(* Logix 5000 project; controller MV vendor 1 type 14 code 217 rev 31.11; software revision 31.00; part 25 of 53 *)
(* tags used below, declared in another part *)
   Alarm_Reset : BOOL;
   comms_to_blunger_write_enabled : BOOL;
   comms_to_fv_route_write_enabled : BOOL;
   comms_to_mv_route_write_enabled : BOOL;
   CWD : CHECKWORD_FLAGS;
   Default_Check_Time : DINT;
   fvrroute_slc_still_active : BOOL;
   Item_Faults_Are_Latched : BOOL;
   Item_Simulation_Flag : BOOL;
   MC_CH2_FM_AI : PlantItem;   // CH2_FM
   mc_comms_from_brewhouse : MESSAGE;
   mc_comms_from_brewhouse_timer : TIMER;
   mc_comms_to_blunger : MESSAGE;
   mc_comms_to_blunger_timer : TIMER;
   mc_comms_to_fv_route : MESSAGE;
   mc_comms_to_fv_route_timer : TIMER;
   mc_comms_to_mv_route : MESSAGE;
   mc_comms_to_mv_route_timer : TIMER;
   MC_N23 : INT[255];   // P2 FLOW Control block and da ta for P2 flowrate P ID loop
   MC_P1 : PlantItem;   // P1
   MC_P1_ALARM : ALARM_DIGITAL;
   MC_P1_D : ALIAS FOR RIO_Rack_2:10:O.Data.0;
   MC_P1_R : ALIAS FOR RIO_Rack_2:11:I.Data.0;
   MC_P1_T : ALIAS FOR RIO_Rack_2:11:I.Data.15;
   MC_P2 : PlantItem;   // P2
   MC_P2_ALARM : ALARM_DIGITAL;
   MC_P2_D : ALIAS FOR RIO_Rack_2:10:O.Data.1;
   MC_P2_Flow_PID : PID;
   MC_P2_R : ALIAS FOR RIO_Rack_2:11:I.Data.1;
   MC_P2_T : ALIAS FOR RIO_Rack_2:11:I.Data.16;
   MC_P3 : PlantItem;   // P3
   MC_P3_ALARM : ALARM_DIGITAL;
   MC_P3_D : ALIAS FOR RIO_Rack_2:10:O.Data.2;
   MC_P3_R : ALIAS FOR RIO_Rack_2:11:I.Data.2;
   MC_P4 : PlantItem;   // P4
   MC_P4_ALARM : ALARM_DIGITAL;
   MC_P4_D : ALIAS FOR RIO_Rack_2:10:O.Data.3;
   MC_P4_R : ALIAS FOR RIO_Rack_2:11:I.Data.3;
   MC_SP_R1_1 : PlantItem;   // SP_R1_1
   MC_SP_R1_1_ALARM : ALARM_DIGITAL;
   MC_SP_R1_1_D : ALIAS FOR RIO_Rack_2:10:O.Data.4;
   MC_SP_R1_1_R : ALIAS FOR RIO_Rack_2:11:I.Data.4;
   MC_SP_R2_1 : PlantItem;   // SP_R2_1
   MC_SP_R2_1_ALARM : ALARM_DIGITAL;
   MC_SP_R2_1_D : ALIAS FOR RIO_Rack_2:10:O.Data.5;
   MC_SP_R2_1_R : ALIAS FOR RIO_Rack_2:11:I.Data.5;
   MC_SP_R2_2 : PlantItem;   // SP_R2_2
   MC_SP_R2_2_ALARM : ALARM_DIGITAL;
   MC_SP_R2_2_D : ALIAS FOR RIO_Rack_2:10:O.Data.15;
   MC_SP_R2_2_R : ALIAS FOR RIO_Rack_2:11:I.Data.14;
   MC_SP_R3_1 : PlantItem;   // SP_R3_1
   MC_SP_R3_1_ALARM : ALARM_DIGITAL;
   MC_SP_R3_1_D : ALIAS FOR RIO_Rack_2:10:O.Data.6;
   MC_SP_R3_1_R : ALIAS FOR RIO_Rack_2:11:I.Data.6;
   MC_SP_R5_1 : PlantItem;   // SP_R5_1
   MC_SP_R5_1_ALARM : ALARM_DIGITAL;
   MC_SP_R5_1_D : ALIAS FOR RIO_Rack_2:10:O.Data.7;
   MC_SP_R5_1_R : ALIAS FOR RIO_Rack_2:11:I.Data.7;
   MC_SP_R5_2 : PlantItem;   // SP_R5_2
   MC_SP_R5_2_ALARM : ALARM_DIGITAL;
   MC_SP_R5_2_D : ALIAS FOR RIO_Rack_2:10:O.Data.8;
   MC_SP_R5_2_R : ALIAS FOR RIO_Rack_2:11:I.Data.8;
   MC_SP_R6_1 : PlantItem;   // SP_R6_1
   MC_SP_R6_1_ALARM : ALARM_DIGITAL;
   MC_SP_R6_1_D : ALIAS FOR RIO_Rack_2:10:O.Data.9;
   MC_SP_R6_1_R : ALIAS FOR RIO_Rack_2:11:I.Data.9;
   MC_SP_R6_2 : PlantItem;   // SP_R6_2
   MC_SP_R6_2_ALARM : ALARM_DIGITAL;
   MC_SP_R6_2_D : ALIAS FOR RIO_Rack_2:10:O.Data.10;
   MC_SP_R6_2_R : ALIAS FOR RIO_Rack_2:11:I.Data.10;
   MC_SP_R6_3 : PlantItem;   // SP_R6_3
   MC_SP_R6_3_ALARM : ALARM_DIGITAL;
   MC_SP_R6_3_D : ALIAS FOR RIO_Rack_2:10:O.Data.11;
   MC_SP_R6_3_R : ALIAS FOR RIO_Rack_2:11:I.Data.11;
   MC_SP_R6_4 : PlantItem;   // SP_R6_4
   MC_SP_R6_4_ALARM : ALARM_DIGITAL;
   MC_SP_R6_4_D : ALIAS FOR RIO_Rack_2:10:O.Data.12;
   MC_SP_R6_4_R : ALIAS FOR RIO_Rack_2:11:I.Data.12;
   MC_SP_R6_5 : PlantItem;   // SP_R6_5
   MC_SP_R6_5_ALARM : ALARM_DIGITAL;
   MC_SP_R6_5_D : ALIAS FOR RIO_Rack_2:10:O.Data.13;
   MC_SP_R6_5_R : ALIAS FOR RIO_Rack_2:11:I.Data.13;
   One_Second_One_Scan : ALIAS FOR One_Second_1_scan;
   reset_msg_interval : BOOL;
   Scada_Pump_Fault_No : DINT;
   Scada_Pump_H_Fault_No : DINT;
   Scada_Pump_T_Fault_No : DINT;
   Unused_Healthy_Feedback : BOOL;
   Unused_NotTripped_Feedback : BOOL;
(* MC_Common, continued *)

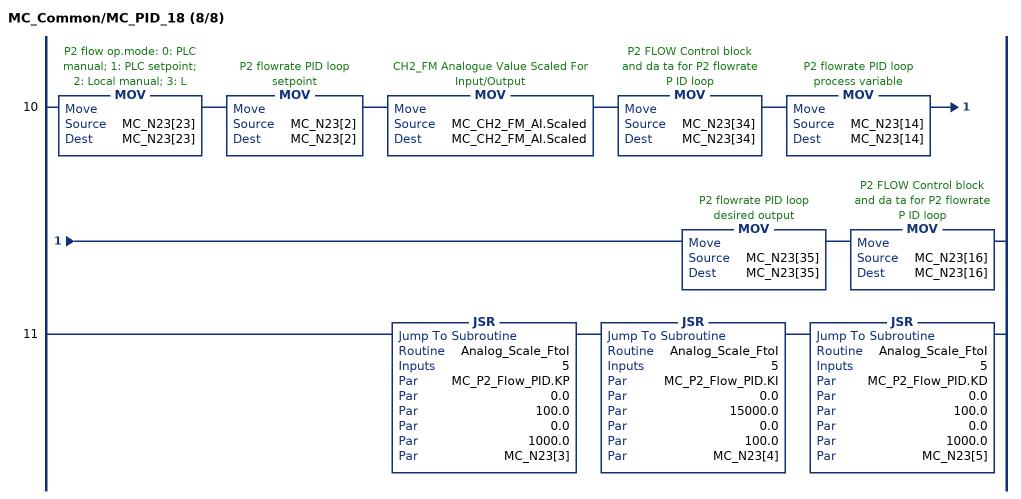
   [picture p462: MC_Common/MC_PID_18 rungs 10-11]
   10: MOV(MC_N23[23],MC_N23[23])MOV(MC_N23[2],MC_N23[2])MOV(MC_CH2_FM_AI.Scaled,MC_CH2_FM_AI.Scaled)MOV(MC_N23[34],MC_N23[34])MOV(MC_N23[14],MC_N23[14])MOV(MC_N23[35],MC_N23[35])MOV(MC_N23[16],MC_N23[16]);
   11: JSR(Analog_Scale_FtoI,5,MC_P2_Flow_PID.KP,0.0,100.0,0.0,1000.0,MC_N23[3])JSR(Analog_Scale_FtoI,5,MC_P2_Flow_PID.KI,0.0,15000.0,0.0,100.0,MC_N23[4])JSR(Analog_Scale_FtoI,5,MC_P2_Flow_PID.KD,0.0,100.0,0.0,1000.0,MC_N23[5]);
END_ROUTINE

ROUTINE MC_PLC_WRITE_REPLACEMENTS   (* ladder *)
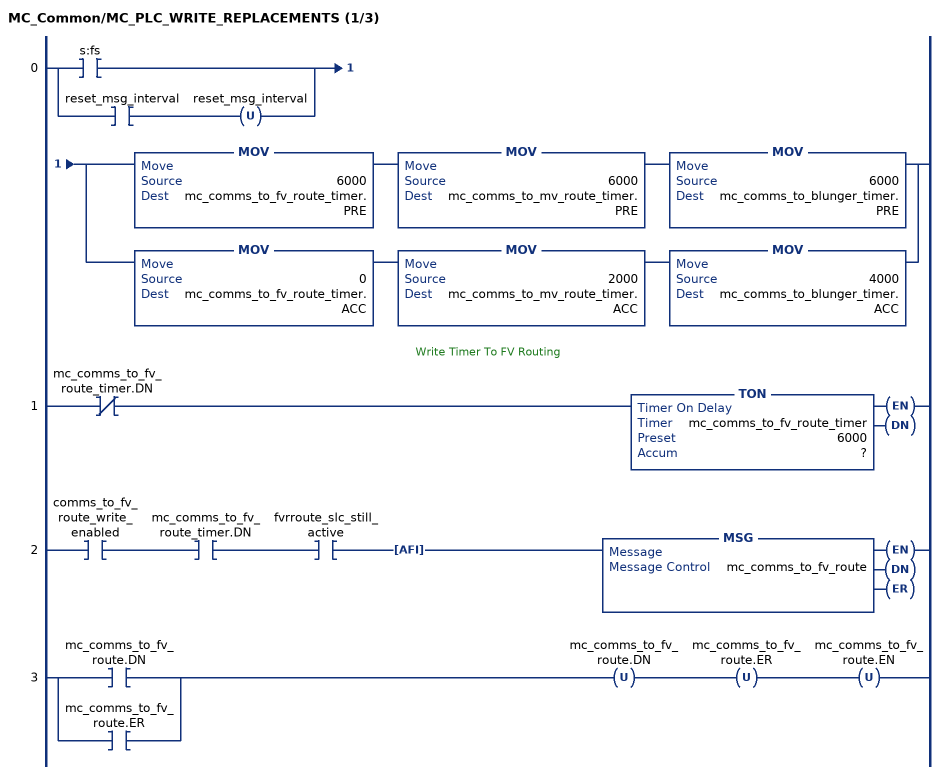
   0: [XIC(s:fs) ,XIC(reset_msg_interval) OTU(reset_msg_interval) ][MOV(6000,mc_comms_to_fv_route_timer.PRE) MOV(6000,mc_comms_to_mv_route_timer.PRE) MOV(6000,mc_comms_to_blunger_timer.PRE) ,MOV(0,mc_comms_to_fv_route_timer.ACC) MOV(2000,mc_comms_to_mv_route_timer.ACC) MOV(4000,mc_comms_to_blunger_timer.ACC) ];
   // Write Timer To FV Routing
   1: XIO(mc_comms_to_fv_route_timer.DN)TON(mc_comms_to_fv_route_timer,?,?);
   2: XIC(comms_to_fv_route_write_enabled)XIC(mc_comms_to_fv_route_timer.DN)XIC(fvrroute_slc_still_active)AFI()MSG(mc_comms_to_fv_route);
   3: [XIC(mc_comms_to_fv_route.DN) ,XIC(mc_comms_to_fv_route.ER) ]OTU(mc_comms_to_fv_route.DN)OTU(mc_comms_to_fv_route.ER)OTU(mc_comms_to_fv_route.EN);
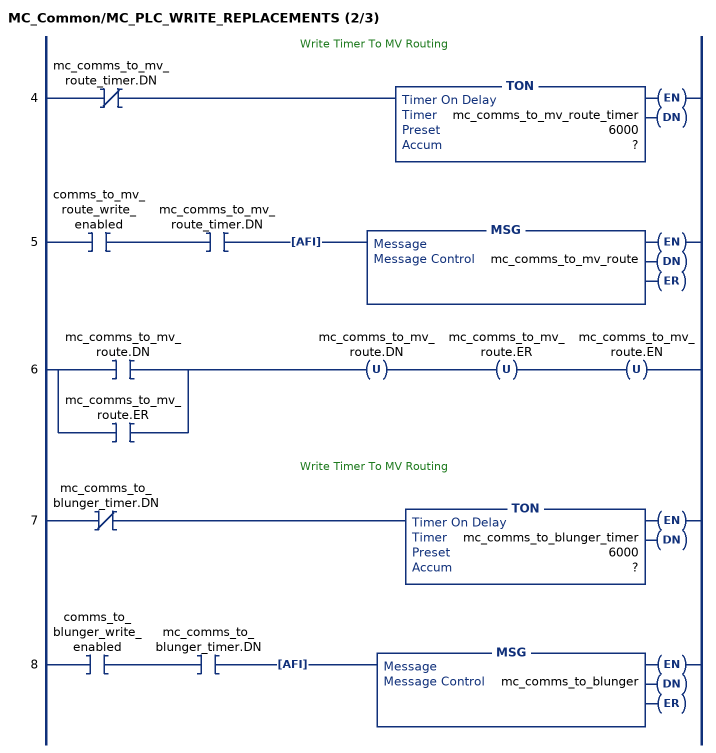
   // Write Timer To MV Routing
   4: XIO(mc_comms_to_mv_route_timer.DN)TON(mc_comms_to_mv_route_timer,?,?);
   5: XIC(comms_to_mv_route_write_enabled)XIC(mc_comms_to_mv_route_timer.DN)AFI()MSG(mc_comms_to_mv_route);
   6: [XIC(mc_comms_to_mv_route.DN) ,XIC(mc_comms_to_mv_route.ER) ]OTU(mc_comms_to_mv_route.DN)OTU(mc_comms_to_mv_route.ER)OTU(mc_comms_to_mv_route.EN);
   // Write Timer To MV Routing
   7: XIO(mc_comms_to_blunger_timer.DN)TON(mc_comms_to_blunger_timer,?,?);
   8: XIC(comms_to_blunger_write_enabled)XIC(mc_comms_to_blunger_timer.DN)AFI()MSG(mc_comms_to_blunger);
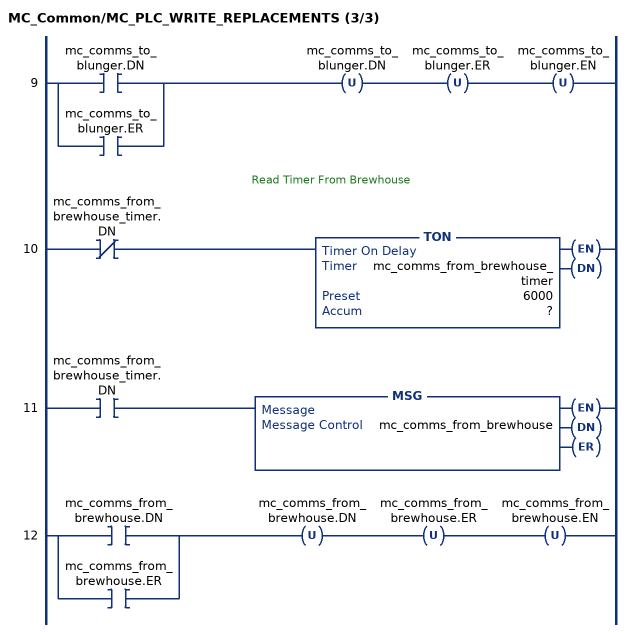
   9: [XIC(mc_comms_to_blunger.DN) ,XIC(mc_comms_to_blunger.ER) ]OTU(mc_comms_to_blunger.DN)OTU(mc_comms_to_blunger.ER)OTU(mc_comms_to_blunger.EN);
   // Read Timer From Brewhouse
   10: XIO(mc_comms_from_brewhouse_timer.DN)TON(mc_comms_from_brewhouse_timer,?,?);
   11: XIC(mc_comms_from_brewhouse_timer.DN)MSG(mc_comms_from_brewhouse);
   12: [XIC(mc_comms_from_brewhouse.DN) ,XIC(mc_comms_from_brewhouse.ER) ]OTU(mc_comms_from_brewhouse.DN)OTU(mc_comms_from_brewhouse.ER)OTU(mc_comms_from_brewhouse.EN);
END_ROUTINE

ROUTINE MC_Pumps   (* ladder *)
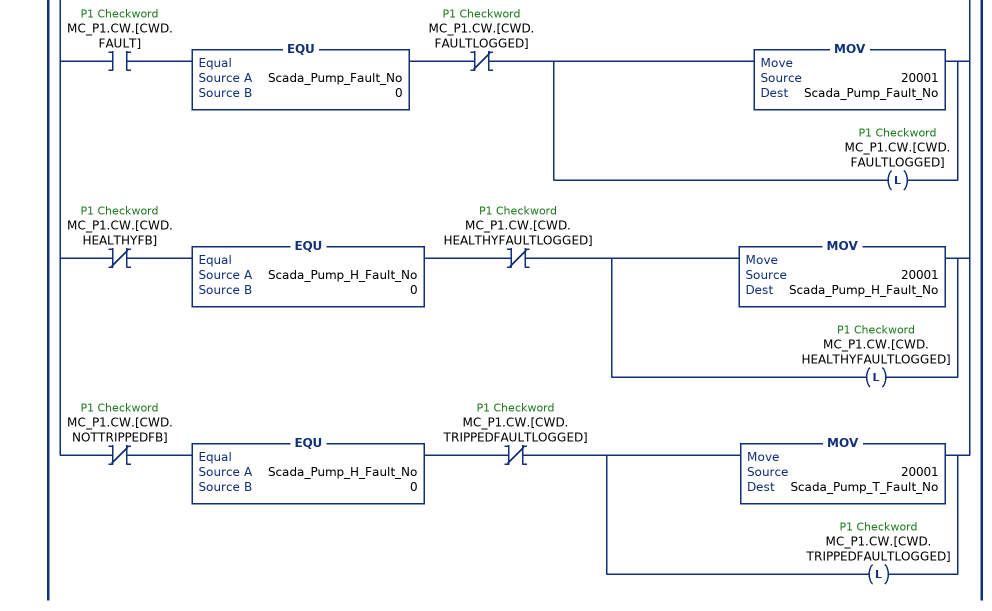
   0: [NEQ(MC_P1.DriveBits,0) OTE(MC_P1.CW.[CWD.AUTODRV]) ,[XIC(MC_P1.CW.[CWD.AUTODRV]) XIO(MC_P1.CW.[CWD.MANUAL]) ,XIC(MC_P1.CW.[CWD.MANDRV]) XIC(MC_P1.CW.[CWD.MANUAL]) ] OTE(MC_P1.CW.[CWD.OUTPUT]) ,XIC(MC_P1.CW.[CWD.OUTPUT]) OTE(MC_P1_D) ,XIC(S:FS) [OTU(MC_P1.CW.[CWD.MANUAL]) ,LEQ(MC_P1.CheckTime,0) MOV(Default_Check_Time,MC_P1.CheckTime) ] ,[[XIC(MC_P1_R) XIO(Item_Simulation_Flag) ,XIC(Item_Simulation_Flag) [XIC(MC_P1.CW.[CWD.OUTPUT]) XIO(MC_P1.CW.[CWD.SIMFAIL]) ,XIO(MC_P1.CW.[CWD.OUTPUT]) XIC(MC_P1.CW.[CWD.SIMFAIL]) ] ] OTE(MC_P1.CW.[CWD.RUNFB]) ,[XIC(Item_Simulation_Flag) ,XIC(MC_P1.CW.[CWD.CHECKOFF]) ,XIC(Unused_Healthy_Feedback) ] OTE(MC_P1.CW.[CWD.HEALTHYFB]) ,[XIC(Item_Simulation_Flag) ,XIC(MC_P1.CW.[CWD.CHECKOFF]) ,XIO(MC_P1_T) ] OTE(MC_P1.CW.[CWD.NOTTRIPPEDFB]) ] ,[XIC(MC_P1.CW.[CWD.OUTPUT]) XIO(MC_P1.CW.[CWD.PREVSCAN]) ,XIO(MC_P1.CW.[CWD.OUTPUT]) XIC(MC_P1.CW.[CWD.PREVSCAN]) ] CLR(MC_P1.CheckTimer) ,XIC(One_Second_One_Scan) LES(MC_P1.CheckTimer,MC_P1.CheckTime) ADD(MC_P1.CheckTimer,1,MC_P1.CheckTimer) ,XIO(MC_P1.CW.[CWD.FAULT]) OTU(MC_P1.CW.[CWD.FAULTLOGGED]) ,[GEQ(MC_P1.CheckTimer,MC_P1.CheckTime) [XIC(MC_P1.CW.[CWD.OUTPUT]) XIO(MC_P1.CW.[CWD.RUNFB]) ,XIO(MC_P1.CW.[CWD.OUTPUT]) XIC(MC_P1.CW.[CWD.RUNFB]) ] ,XIO(MC_P1.CW.[CWD.HEALTHYFB]) ,XIO(MC_P1.CW.[CWD.NOTTRIPPEDFB]) ,XIC(MC_P1.CW.[CWD.FAULT]) XIC(Item_Faults_Are_Latched) ,XIC(MC_P1.CW.[CWD.HIGHLIGHT]) ] XIO(MC_P1.CW.[CWD.CHECKOFF]) XIO(Alarm_Reset) [OTE(MC_P1.CW.[CWD.FAULT]) ,ALMD(MC_P1_ALARM,0,0,0,0) ] ,XIC(MC_P1.CW.[CWD.OUTPUT]) OTE(MC_P1.CW.[CWD.PREVSCAN]) ,XIC(MC_P1.CW.[CWD.FAULT]) EQU(Scada_Pump_Fault_No,0) XIO(MC_P1.CW.[CWD.FAULTLOGGED]) [MOV(20001,Scada_Pump_Fault_No) ,OTL(MC_P1.CW.[CWD.FAULTLOGGED]) ] ,XIO(MC_P1.CW.[CWD.HEALTHYFB]) EQU(Scada_Pump_H_Fault_No,0) XIO(MC_P1.CW.[CWD.HEALTHYFAULTLOGGED]) [MOV(20001,Scada_Pump_H_Fault_No) ,OTL(MC_P1.CW.[CWD.HEALTHYFAULTLOGGED]) ] ,XIO(MC_P1.CW.[CWD.NOTTRIPPEDFB]) EQU(Scada_Pump_H_Fault_No,0) XIO(MC_P1.CW.[CWD.TRIPPEDFAULTLOGGED]) [MOV(20001,Scada_Pump_T_Fault_No) ,OTL(MC_P1.CW.[CWD.TRIPPEDFAULTLOGGED]) ] ];
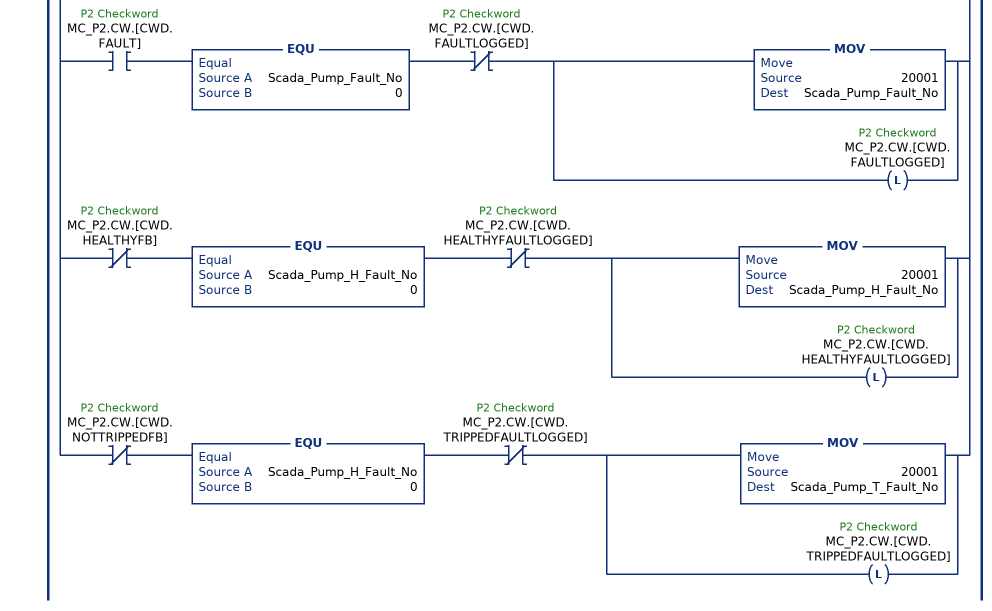
   1: [NEQ(MC_P2.DriveBits,0) OTE(MC_P2.CW.[CWD.AUTODRV]) ,[XIC(MC_P2.CW.[CWD.AUTODRV]) XIO(MC_P2.CW.[CWD.MANUAL]) ,XIC(MC_P2.CW.[CWD.MANDRV]) XIC(MC_P2.CW.[CWD.MANUAL]) ] OTE(MC_P2.CW.[CWD.OUTPUT]) ,XIC(MC_P2.CW.[CWD.OUTPUT]) OTE(MC_P2_D) ,XIC(S:FS) [OTU(MC_P2.CW.[CWD.MANUAL]) ,LEQ(MC_P2.CheckTime,0) MOV(Default_Check_Time,MC_P2.CheckTime) ] ,[[XIC(MC_P2_R) XIO(Item_Simulation_Flag) ,XIC(Item_Simulation_Flag) [XIC(MC_P2.CW.[CWD.OUTPUT]) XIO(MC_P2.CW.[CWD.SIMFAIL]) ,XIO(MC_P2.CW.[CWD.OUTPUT]) XIC(MC_P2.CW.[CWD.SIMFAIL]) ] ] OTE(MC_P2.CW.[CWD.RUNFB]) ,[XIC(Item_Simulation_Flag) ,XIC(MC_P2.CW.[CWD.CHECKOFF]) ,XIC(Unused_Healthy_Feedback) ] OTE(MC_P2.CW.[CWD.HEALTHYFB]) ,[XIC(Item_Simulation_Flag) ,XIC(MC_P2.CW.[CWD.CHECKOFF]) ,XIC(MC_P2_T) ] OTE(MC_P2.CW.[CWD.NOTTRIPPEDFB]) ] ,[XIC(MC_P2.CW.[CWD.OUTPUT]) XIO(MC_P2.CW.[CWD.PREVSCAN]) ,XIO(MC_P2.CW.[CWD.OUTPUT]) XIC(MC_P2.CW.[CWD.PREVSCAN]) ] CLR(MC_P2.CheckTimer) ,XIC(One_Second_One_Scan) LES(MC_P2.CheckTimer,MC_P2.CheckTime) ADD(MC_P2.CheckTimer,1,MC_P2.CheckTimer) ,XIO(MC_P2.CW.[CWD.FAULT]) OTU(MC_P2.CW.[CWD.FAULTLOGGED]) ,[GEQ(MC_P2.CheckTimer,MC_P2.CheckTime) [XIC(MC_P2.CW.[CWD.OUTPUT]) XIO(MC_P2.CW.[CWD.RUNFB]) ,XIO(MC_P2.CW.[CWD.OUTPUT]) XIC(MC_P2.CW.[CWD.RUNFB]) ] ,XIO(MC_P2.CW.[CWD.HEALTHYFB]) ,XIO(MC_P2.CW.[CWD.NOTTRIPPEDFB]) ,XIC(MC_P2.CW.[CWD.FAULT]) XIC(Item_Faults_Are_Latched) ,XIC(MC_P2.CW.[CWD.HIGHLIGHT]) ] XIO(MC_P2.CW.[CWD.CHECKOFF]) XIO(Alarm_Reset) [OTE(MC_P2.CW.[CWD.FAULT]) ,ALMD(MC_P2_ALARM,0,0,0,0) ] ,XIC(MC_P2.CW.[CWD.OUTPUT]) OTE(MC_P2.CW.[CWD.PREVSCAN]) ,XIC(MC_P2.CW.[CWD.FAULT]) EQU(Scada_Pump_Fault_No,0) XIO(MC_P2.CW.[CWD.FAULTLOGGED]) [MOV(20001,Scada_Pump_Fault_No) ,OTL(MC_P2.CW.[CWD.FAULTLOGGED]) ] ,XIO(MC_P2.CW.[CWD.HEALTHYFB]) EQU(Scada_Pump_H_Fault_No,0) XIO(MC_P2.CW.[CWD.HEALTHYFAULTLOGGED]) [MOV(20001,Scada_Pump_H_Fault_No) ,OTL(MC_P2.CW.[CWD.HEALTHYFAULTLOGGED]) ] ,XIO(MC_P2.CW.[CWD.NOTTRIPPEDFB]) EQU(Scada_Pump_H_Fault_No,0) XIO(MC_P2.CW.[CWD.TRIPPEDFAULTLOGGED]) [MOV(20001,Scada_Pump_T_Fault_No) ,OTL(MC_P2.CW.[CWD.TRIPPEDFAULTLOGGED]) ] ];
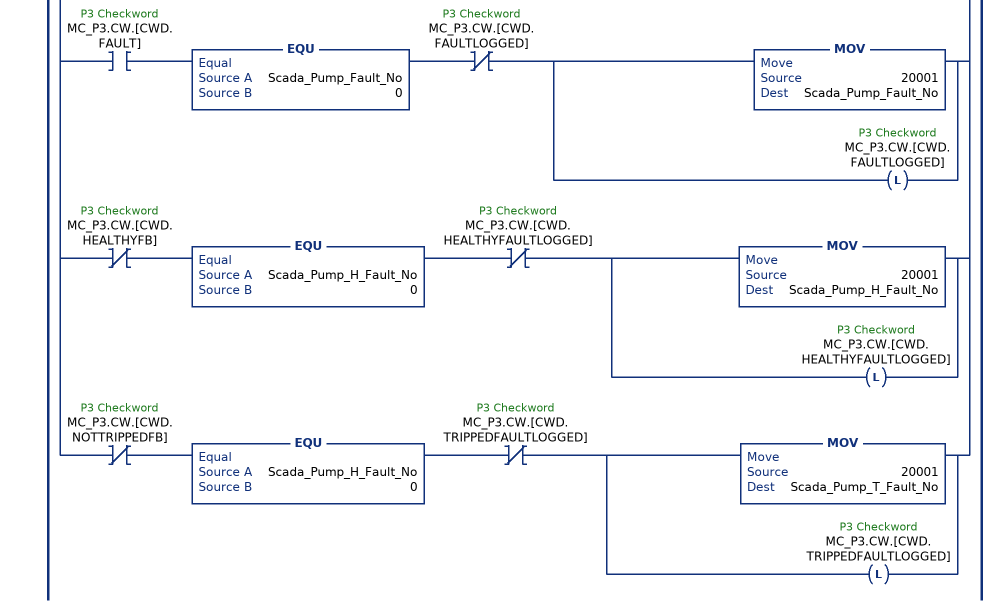
   2: [NEQ(MC_P3.DriveBits,0) OTE(MC_P3.CW.[CWD.AUTODRV]) ,[XIC(MC_P3.CW.[CWD.AUTODRV]) XIO(MC_P3.CW.[CWD.MANUAL]) ,XIC(MC_P3.CW.[CWD.MANDRV]) XIC(MC_P3.CW.[CWD.MANUAL]) ] OTE(MC_P3.CW.[CWD.OUTPUT]) ,XIC(MC_P3.CW.[CWD.OUTPUT]) OTE(MC_P3_D) ,XIC(S:FS) [OTU(MC_P3.CW.[CWD.MANUAL]) ,LEQ(MC_P3.CheckTime,0) MOV(Default_Check_Time,MC_P3.CheckTime) ] ,[[XIC(MC_P3_R) XIO(Item_Simulation_Flag) ,XIC(Item_Simulation_Flag) [XIC(MC_P3.CW.[CWD.OUTPUT]) XIO(MC_P3.CW.[CWD.SIMFAIL]) ,XIO(MC_P3.CW.[CWD.OUTPUT]) XIC(MC_P3.CW.[CWD.SIMFAIL]) ] ] OTE(MC_P3.CW.[CWD.RUNFB]) ,[XIC(Item_Simulation_Flag) ,XIC(MC_P3.CW.[CWD.CHECKOFF]) ,XIC(Unused_Healthy_Feedback) ] OTE(MC_P3.CW.[CWD.HEALTHYFB]) ,[XIC(Item_Simulation_Flag) ,XIC(MC_P3.CW.[CWD.CHECKOFF]) ,XIC(Unused_NotTripped_Feedback) ] OTE(MC_P3.CW.[CWD.NOTTRIPPEDFB]) ] ,[XIC(MC_P3.CW.[CWD.OUTPUT]) XIO(MC_P3.CW.[CWD.PREVSCAN]) ,XIO(MC_P3.CW.[CWD.OUTPUT]) XIC(MC_P3.CW.[CWD.PREVSCAN]) ] CLR(MC_P3.CheckTimer) ,XIC(One_Second_One_Scan) LES(MC_P3.CheckTimer,MC_P3.CheckTime) ADD(MC_P3.CheckTimer,1,MC_P3.CheckTimer) ,XIO(MC_P3.CW.[CWD.FAULT]) OTU(MC_P3.CW.[CWD.FAULTLOGGED]) ,[GEQ(MC_P3.CheckTimer,MC_P3.CheckTime) [XIC(MC_P3.CW.[CWD.OUTPUT]) XIO(MC_P3.CW.[CWD.RUNFB]) ,XIO(MC_P3.CW.[CWD.OUTPUT]) XIC(MC_P3.CW.[CWD.RUNFB]) ] ,XIO(MC_P3.CW.[CWD.HEALTHYFB]) ,XIO(MC_P3.CW.[CWD.NOTTRIPPEDFB]) ,XIC(MC_P3.CW.[CWD.FAULT]) XIC(Item_Faults_Are_Latched) ,XIC(MC_P3.CW.[CWD.HIGHLIGHT]) ] XIO(MC_P3.CW.[CWD.CHECKOFF]) XIO(Alarm_Reset) [OTE(MC_P3.CW.[CWD.FAULT]) ,ALMD(MC_P3_ALARM,0,0,0,0) ] ,XIC(MC_P3.CW.[CWD.OUTPUT]) OTE(MC_P3.CW.[CWD.PREVSCAN]) ,XIC(MC_P3.CW.[CWD.FAULT]) EQU(Scada_Pump_Fault_No,0) XIO(MC_P3.CW.[CWD.FAULTLOGGED]) [MOV(20001,Scada_Pump_Fault_No) ,OTL(MC_P3.CW.[CWD.FAULTLOGGED]) ] ,XIO(MC_P3.CW.[CWD.HEALTHYFB]) EQU(Scada_Pump_H_Fault_No,0) XIO(MC_P3.CW.[CWD.HEALTHYFAULTLOGGED]) [MOV(20001,Scada_Pump_H_Fault_No) ,OTL(MC_P3.CW.[CWD.HEALTHYFAULTLOGGED]) ] ,XIO(MC_P3.CW.[CWD.NOTTRIPPEDFB]) EQU(Scada_Pump_H_Fault_No,0) XIO(MC_P3.CW.[CWD.TRIPPEDFAULTLOGGED]) [MOV(20001,Scada_Pump_T_Fault_No) ,OTL(MC_P3.CW.[CWD.TRIPPEDFAULTLOGGED]) ] ];
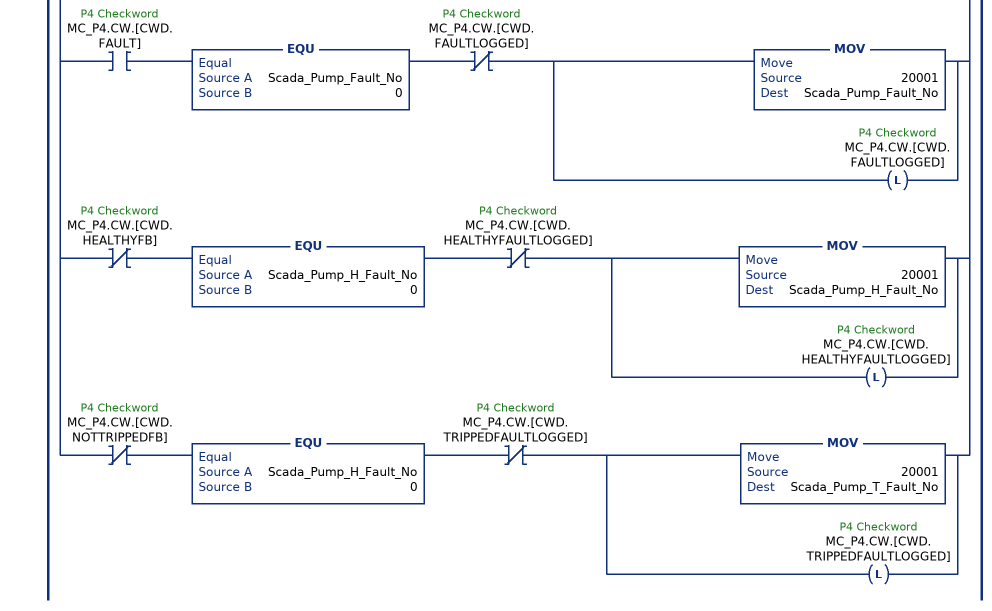
   3: [NEQ(MC_P4.DriveBits,0) OTE(MC_P4.CW.[CWD.AUTODRV]) ,[XIC(MC_P4.CW.[CWD.AUTODRV]) XIO(MC_P4.CW.[CWD.MANUAL]) ,XIC(MC_P4.CW.[CWD.MANDRV]) XIC(MC_P4.CW.[CWD.MANUAL]) ] OTE(MC_P4.CW.[CWD.OUTPUT]) ,XIC(MC_P4.CW.[CWD.OUTPUT]) OTE(MC_P4_D) ,XIC(S:FS) [OTU(MC_P4.CW.[CWD.MANUAL]) ,LEQ(MC_P4.CheckTime,0) MOV(Default_Check_Time,MC_P4.CheckTime) ] ,[[XIC(MC_P4_R) XIO(Item_Simulation_Flag) ,XIC(Item_Simulation_Flag) [XIC(MC_P4.CW.[CWD.OUTPUT]) XIO(MC_P4.CW.[CWD.SIMFAIL]) ,XIO(MC_P4.CW.[CWD.OUTPUT]) XIC(MC_P4.CW.[CWD.SIMFAIL]) ] ] OTE(MC_P4.CW.[CWD.RUNFB]) ,[XIC(Item_Simulation_Flag) ,XIC(MC_P4.CW.[CWD.CHECKOFF]) ,XIC(Unused_Healthy_Feedback) ] OTE(MC_P4.CW.[CWD.HEALTHYFB]) ,[XIC(Item_Simulation_Flag) ,XIC(MC_P4.CW.[CWD.CHECKOFF]) ,XIC(Unused_NotTripped_Feedback) ] OTE(MC_P4.CW.[CWD.NOTTRIPPEDFB]) ] ,[XIC(MC_P4.CW.[CWD.OUTPUT]) XIO(MC_P4.CW.[CWD.PREVSCAN]) ,XIO(MC_P4.CW.[CWD.OUTPUT]) XIC(MC_P4.CW.[CWD.PREVSCAN]) ] CLR(MC_P4.CheckTimer) ,XIC(One_Second_One_Scan) LES(MC_P4.CheckTimer,MC_P4.CheckTime) ADD(MC_P4.CheckTimer,1,MC_P4.CheckTimer) ,XIO(MC_P4.CW.[CWD.FAULT]) OTU(MC_P4.CW.[CWD.FAULTLOGGED]) ,[GEQ(MC_P4.CheckTimer,MC_P4.CheckTime) [XIC(MC_P4.CW.[CWD.OUTPUT]) XIO(MC_P4.CW.[CWD.RUNFB]) ,XIO(MC_P4.CW.[CWD.OUTPUT]) XIC(MC_P4.CW.[CWD.RUNFB]) ] ,XIO(MC_P4.CW.[CWD.HEALTHYFB]) ,XIO(MC_P4.CW.[CWD.NOTTRIPPEDFB]) ,XIC(MC_P4.CW.[CWD.FAULT]) XIC(Item_Faults_Are_Latched) ,XIC(MC_P4.CW.[CWD.HIGHLIGHT]) ] XIO(MC_P4.CW.[CWD.CHECKOFF]) XIO(Alarm_Reset) [OTE(MC_P4.CW.[CWD.FAULT]) ,ALMD(MC_P4_ALARM,0,0,0,0) ] ,XIC(MC_P4.CW.[CWD.OUTPUT]) OTE(MC_P4.CW.[CWD.PREVSCAN]) ,XIC(MC_P4.CW.[CWD.FAULT]) EQU(Scada_Pump_Fault_No,0) XIO(MC_P4.CW.[CWD.FAULTLOGGED]) [MOV(20001,Scada_Pump_Fault_No) ,OTL(MC_P4.CW.[CWD.FAULTLOGGED]) ] ,XIO(MC_P4.CW.[CWD.HEALTHYFB]) EQU(Scada_Pump_H_Fault_No,0) XIO(MC_P4.CW.[CWD.HEALTHYFAULTLOGGED]) [MOV(20001,Scada_Pump_H_Fault_No) ,OTL(MC_P4.CW.[CWD.HEALTHYFAULTLOGGED]) ] ,XIO(MC_P4.CW.[CWD.NOTTRIPPEDFB]) EQU(Scada_Pump_H_Fault_No,0) XIO(MC_P4.CW.[CWD.TRIPPEDFAULTLOGGED]) [MOV(20001,Scada_Pump_T_Fault_No) ,OTL(MC_P4.CW.[CWD.TRIPPEDFAULTLOGGED]) ] ];
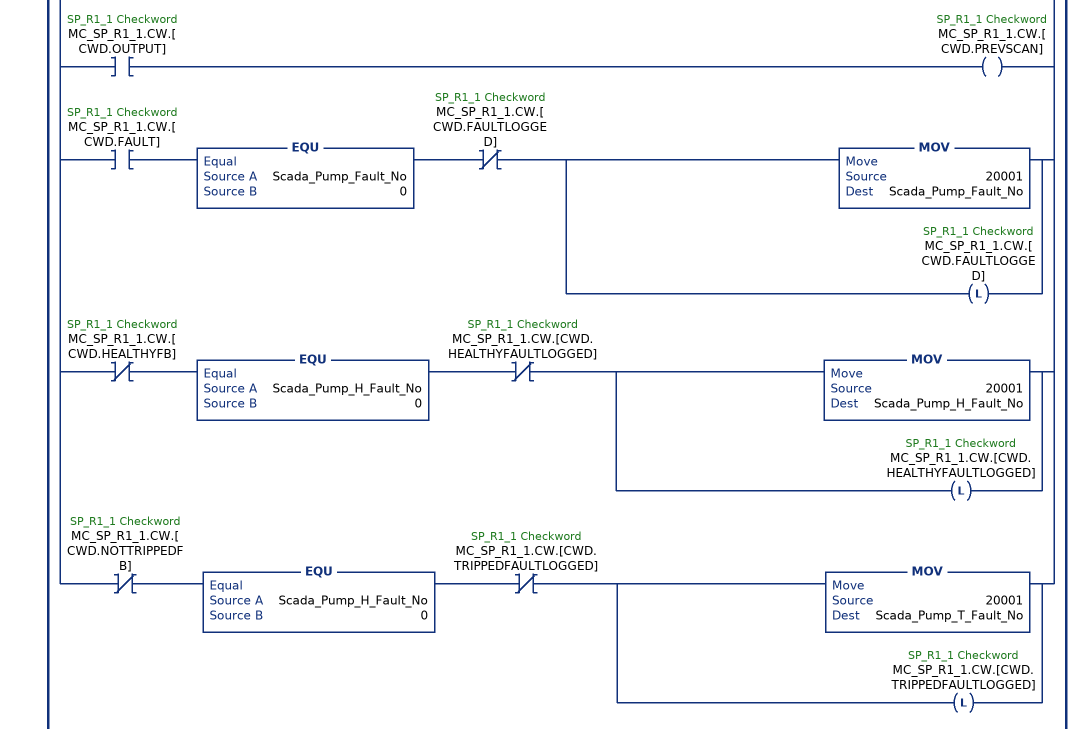
   4: [NEQ(MC_SP_R1_1.DriveBits,0) OTE(MC_SP_R1_1.CW.[CWD.AUTODRV]) ,[XIC(MC_SP_R1_1.CW.[CWD.AUTODRV]) XIO(MC_SP_R1_1.CW.[CWD.MANUAL]) ,XIC(MC_SP_R1_1.CW.[CWD.MANDRV]) XIC(MC_SP_R1_1.CW.[CWD.MANUAL]) ] OTE(MC_SP_R1_1.CW.[CWD.OUTPUT]) ,XIC(MC_SP_R1_1.CW.[CWD.OUTPUT]) OTE(MC_SP_R1_1_D) ,XIC(S:FS) [OTU(MC_SP_R1_1.CW.[CWD.MANUAL]) ,LEQ(MC_SP_R1_1.CheckTime,0) MOV(Default_Check_Time,MC_SP_R1_1.CheckTime) ] ,[[XIC(MC_SP_R1_1_R) XIO(Item_Simulation_Flag) ,XIC(Item_Simulation_Flag) [XIC(MC_SP_R1_1.CW.[CWD.OUTPUT]) XIO(MC_SP_R1_1.CW.[CWD.SIMFAIL]) ,XIO(MC_SP_R1_1.CW.[CWD.OUTPUT]) XIC(MC_SP_R1_1.CW.[CWD.SIMFAIL]) ] ] OTE(MC_SP_R1_1.CW.[CWD.RUNFB]) ,[XIC(Item_Simulation_Flag) ,XIC(MC_SP_R1_1.CW.[CWD.CHECKOFF]) ,XIC(Unused_Healthy_Feedback) ] OTE(MC_SP_R1_1.CW.[CWD.HEALTHYFB]) ,[XIC(Item_Simulation_Flag) ,XIC(MC_SP_R1_1.CW.[CWD.CHECKOFF]) ,XIC(Unused_NotTripped_Feedback) ] OTE(MC_SP_R1_1.CW.[CWD.NOTTRIPPEDFB]) ] ,[XIC(MC_SP_R1_1.CW.[CWD.OUTPUT]) XIO(MC_SP_R1_1.CW.[CWD.PREVSCAN]) ,XIO(MC_SP_R1_1.CW.[CWD.OUTPUT]) XIC(MC_SP_R1_1.CW.[CWD.PREVSCAN]) ] CLR(MC_SP_R1_1.CheckTimer) ,XIC(One_Second_One_Scan) LES(MC_SP_R1_1.CheckTimer,MC_SP_R1_1.CheckTime) ADD(MC_SP_R1_1.CheckTimer,1,MC_SP_R1_1.CheckTimer) ,XIO(MC_SP_R1_1.CW.[CWD.FAULT]) OTU(MC_SP_R1_1.CW.[CWD.FAULTLOGGED]) ,[GEQ(MC_SP_R1_1.CheckTimer,MC_SP_R1_1.CheckTime) [XIC(MC_SP_R1_1.CW.[CWD.OUTPUT]) XIO(MC_SP_R1_1.CW.[CWD.RUNFB]) ,XIO(MC_SP_R1_1.CW.[CWD.OUTPUT]) XIC(MC_SP_R1_1.CW.[CWD.RUNFB]) ] ,XIO(MC_SP_R1_1.CW.[CWD.HEALTHYFB]) ,XIO(MC_SP_R1_1.CW.[CWD.NOTTRIPPEDFB]) ,XIC(MC_SP_R1_1.CW.[CWD.FAULT]) XIC(Item_Faults_Are_Latched) ,XIC(MC_SP_R1_1.CW.[CWD.HIGHLIGHT]) ] XIO(MC_SP_R1_1.CW.[CWD.CHECKOFF]) XIO(Alarm_Reset) [OTE(MC_SP_R1_1.CW.[CWD.FAULT]) ,ALMD(MC_SP_R1_1_ALARM,0,0,0,0) ] ,XIC(MC_SP_R1_1.CW.[CWD.OUTPUT]) OTE(MC_SP_R1_1.CW.[CWD.PREVSCAN]) ,XIC(MC_SP_R1_1.CW.[CWD.FAULT]) EQU(Scada_Pump_Fault_No,0) XIO(MC_SP_R1_1.CW.[CWD.FAULTLOGGED]) [MOV(20001,Scada_Pump_Fault_No) ,OTL(MC_SP_R1_1.CW.[CWD.FAULTLOGGED]) ] ,XIO(MC_SP_R1_1.CW.[CWD.HEALTHYFB]) EQU(Scada_Pump_H_Fault_No,0) XIO(MC_SP_R1_1.CW.[CWD.HEALTHYFAULTLOGGED]) [MOV(20001,Scada_Pump_H_Fault_No) ,OTL(MC_SP_R1_1.CW.[CWD.HEALTHYFAULTLOGGED]) ] ,XIO(MC_SP_R1_1.CW.[CWD.NOTTRIPPEDFB]) EQU(Scada_Pump_H_Fault_No,0) XIO(MC_SP_R1_1.CW.[CWD.TRIPPEDFAULTLOGGED]) [MOV(20001,Scada_Pump_T_Fault_No) ,OTL(MC_SP_R1_1.CW.[CWD.TRIPPEDFAULTLOGGED]) ] ];
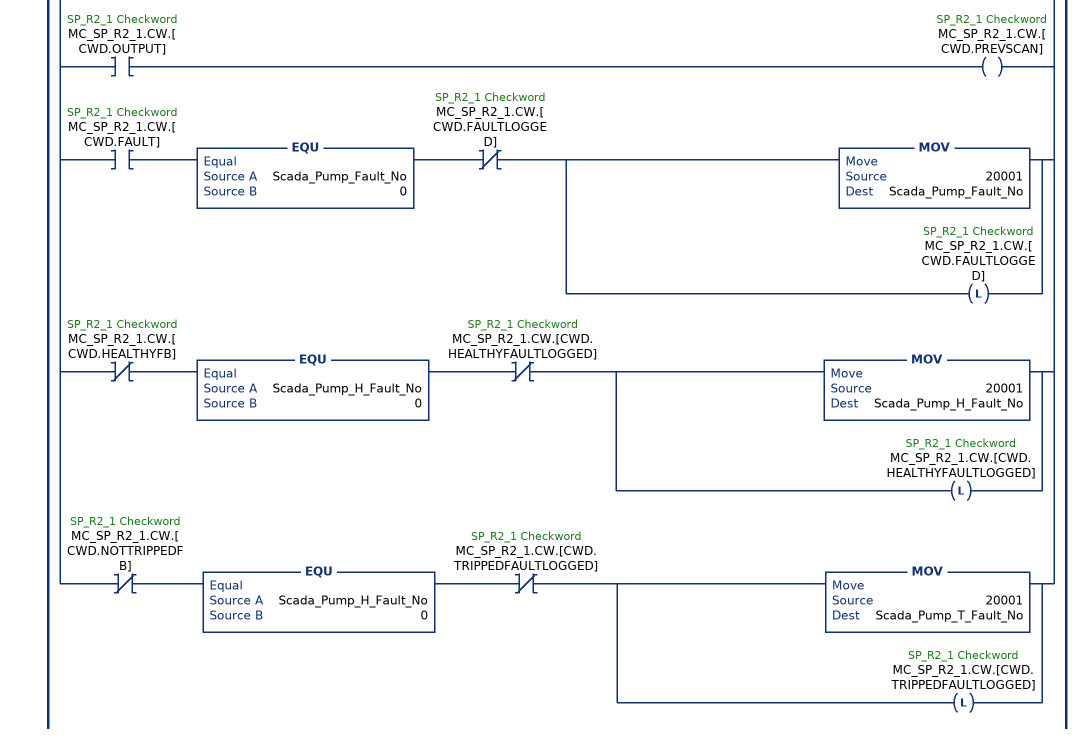
   5: [NEQ(MC_SP_R2_1.DriveBits,0) OTE(MC_SP_R2_1.CW.[CWD.AUTODRV]) ,[XIC(MC_SP_R2_1.CW.[CWD.AUTODRV]) XIO(MC_SP_R2_1.CW.[CWD.MANUAL]) ,XIC(MC_SP_R2_1.CW.[CWD.MANDRV]) XIC(MC_SP_R2_1.CW.[CWD.MANUAL]) ] OTE(MC_SP_R2_1.CW.[CWD.OUTPUT]) ,XIC(MC_SP_R2_1.CW.[CWD.OUTPUT]) OTE(MC_SP_R2_1_D) ,XIC(S:FS) [OTU(MC_SP_R2_1.CW.[CWD.MANUAL]) ,LEQ(MC_SP_R2_1.CheckTime,0) MOV(Default_Check_Time,MC_SP_R2_1.CheckTime) ] ,[[XIC(MC_SP_R2_1_R) XIO(Item_Simulation_Flag) ,XIC(Item_Simulation_Flag) [XIC(MC_SP_R2_1.CW.[CWD.OUTPUT]) XIO(MC_SP_R2_1.CW.[CWD.SIMFAIL]) ,XIO(MC_SP_R2_1.CW.[CWD.OUTPUT]) XIC(MC_SP_R2_1.CW.[CWD.SIMFAIL]) ] ] OTE(MC_SP_R2_1.CW.[CWD.RUNFB]) ,[XIC(Item_Simulation_Flag) ,XIC(MC_SP_R2_1.CW.[CWD.CHECKOFF]) ,XIC(Unused_Healthy_Feedback) ] OTE(MC_SP_R2_1.CW.[CWD.HEALTHYFB]) ,[XIC(Item_Simulation_Flag) ,XIC(MC_SP_R2_1.CW.[CWD.CHECKOFF]) ,XIC(Unused_NotTripped_Feedback) ] OTE(MC_SP_R2_1.CW.[CWD.NOTTRIPPEDFB]) ] ,[XIC(MC_SP_R2_1.CW.[CWD.OUTPUT]) XIO(MC_SP_R2_1.CW.[CWD.PREVSCAN]) ,XIO(MC_SP_R2_1.CW.[CWD.OUTPUT]) XIC(MC_SP_R2_1.CW.[CWD.PREVSCAN]) ] CLR(MC_SP_R2_1.CheckTimer) ,XIC(One_Second_One_Scan) LES(MC_SP_R2_1.CheckTimer,MC_SP_R2_1.CheckTime) ADD(MC_SP_R2_1.CheckTimer,1,MC_SP_R2_1.CheckTimer) ,XIO(MC_SP_R2_1.CW.[CWD.FAULT]) OTU(MC_SP_R2_1.CW.[CWD.FAULTLOGGED]) ,[GEQ(MC_SP_R2_1.CheckTimer,MC_SP_R2_1.CheckTime) [XIC(MC_SP_R2_1.CW.[CWD.OUTPUT]) XIO(MC_SP_R2_1.CW.[CWD.RUNFB]) ,XIO(MC_SP_R2_1.CW.[CWD.OUTPUT]) XIC(MC_SP_R2_1.CW.[CWD.RUNFB]) ] ,XIO(MC_SP_R2_1.CW.[CWD.HEALTHYFB]) ,XIO(MC_SP_R2_1.CW.[CWD.NOTTRIPPEDFB]) ,XIC(MC_SP_R2_1.CW.[CWD.FAULT]) XIC(Item_Faults_Are_Latched) ,XIC(MC_SP_R2_1.CW.[CWD.HIGHLIGHT]) ] XIO(MC_SP_R2_1.CW.[CWD.CHECKOFF]) XIO(Alarm_Reset) [OTE(MC_SP_R2_1.CW.[CWD.FAULT]) ,ALMD(MC_SP_R2_1_ALARM,0,0,0,0) ] ,XIC(MC_SP_R2_1.CW.[CWD.OUTPUT]) OTE(MC_SP_R2_1.CW.[CWD.PREVSCAN]) ,XIC(MC_SP_R2_1.CW.[CWD.FAULT]) EQU(Scada_Pump_Fault_No,0) XIO(MC_SP_R2_1.CW.[CWD.FAULTLOGGED]) [MOV(20001,Scada_Pump_Fault_No) ,OTL(MC_SP_R2_1.CW.[CWD.FAULTLOGGED]) ] ,XIO(MC_SP_R2_1.CW.[CWD.HEALTHYFB]) EQU(Scada_Pump_H_Fault_No,0) XIO(MC_SP_R2_1.CW.[CWD.HEALTHYFAULTLOGGED]) [MOV(20001,Scada_Pump_H_Fault_No) ,OTL(MC_SP_R2_1.CW.[CWD.HEALTHYFAULTLOGGED]) ] ,XIO(MC_SP_R2_1.CW.[CWD.NOTTRIPPEDFB]) EQU(Scada_Pump_H_Fault_No,0) XIO(MC_SP_R2_1.CW.[CWD.TRIPPEDFAULTLOGGED]) [MOV(20001,Scada_Pump_T_Fault_No) ,OTL(MC_SP_R2_1.CW.[CWD.TRIPPEDFAULTLOGGED]) ] ];
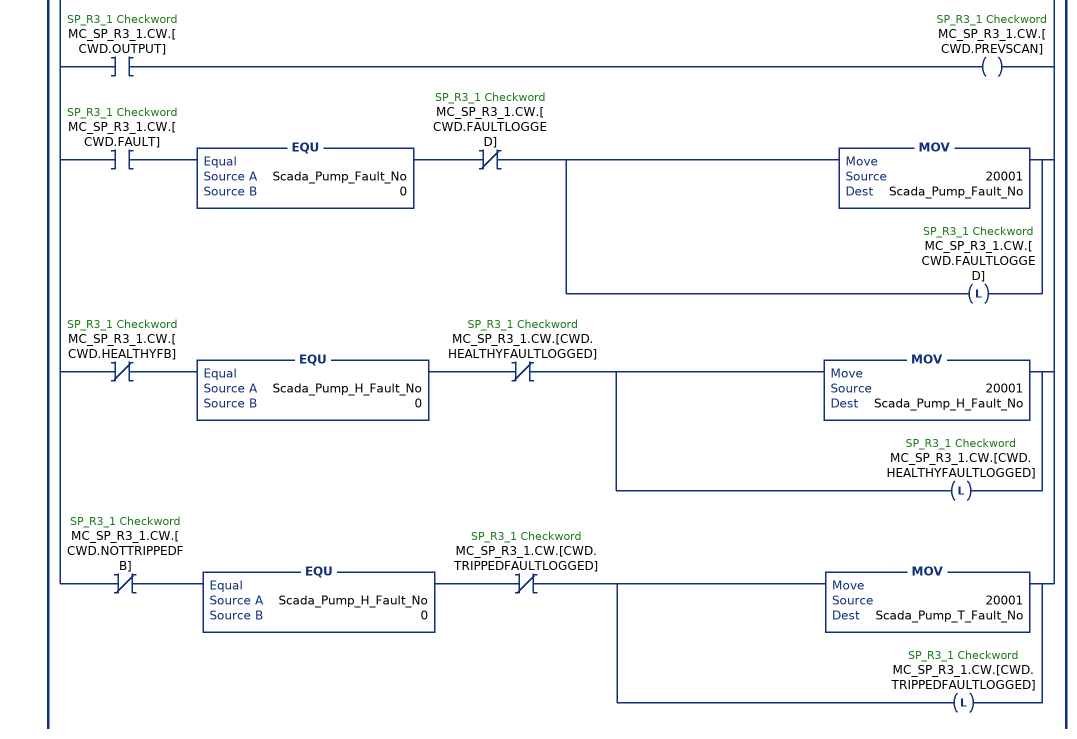
   6: [NEQ(MC_SP_R3_1.DriveBits,0) OTE(MC_SP_R3_1.CW.[CWD.AUTODRV]) ,[XIC(MC_SP_R3_1.CW.[CWD.AUTODRV]) XIO(MC_SP_R3_1.CW.[CWD.MANUAL]) ,XIC(MC_SP_R3_1.CW.[CWD.MANDRV]) XIC(MC_SP_R3_1.CW.[CWD.MANUAL]) ] OTE(MC_SP_R3_1.CW.[CWD.OUTPUT]) ,XIC(MC_SP_R3_1.CW.[CWD.OUTPUT]) OTE(MC_SP_R3_1_D) ,XIC(S:FS) [OTU(MC_SP_R3_1.CW.[CWD.MANUAL]) ,LEQ(MC_SP_R3_1.CheckTime,0) MOV(Default_Check_Time,MC_SP_R3_1.CheckTime) ] ,[[XIC(MC_SP_R3_1_R) XIO(Item_Simulation_Flag) ,XIC(Item_Simulation_Flag) [XIC(MC_SP_R3_1.CW.[CWD.OUTPUT]) XIO(MC_SP_R3_1.CW.[CWD.SIMFAIL]) ,XIO(MC_SP_R3_1.CW.[CWD.OUTPUT]) XIC(MC_SP_R3_1.CW.[CWD.SIMFAIL]) ] ] OTE(MC_SP_R3_1.CW.[CWD.RUNFB]) ,[XIC(Item_Simulation_Flag) ,XIC(MC_SP_R3_1.CW.[CWD.CHECKOFF]) ,XIC(Unused_Healthy_Feedback) ] OTE(MC_SP_R3_1.CW.[CWD.HEALTHYFB]) ,[XIC(Item_Simulation_Flag) ,XIC(MC_SP_R3_1.CW.[CWD.CHECKOFF]) ,XIC(Unused_NotTripped_Feedback) ] OTE(MC_SP_R3_1.CW.[CWD.NOTTRIPPEDFB]) ] ,[XIC(MC_SP_R3_1.CW.[CWD.OUTPUT]) XIO(MC_SP_R3_1.CW.[CWD.PREVSCAN]) ,XIO(MC_SP_R3_1.CW.[CWD.OUTPUT]) XIC(MC_SP_R3_1.CW.[CWD.PREVSCAN]) ] CLR(MC_SP_R3_1.CheckTimer) ,XIC(One_Second_One_Scan) LES(MC_SP_R3_1.CheckTimer,MC_SP_R3_1.CheckTime) ADD(MC_SP_R3_1.CheckTimer,1,MC_SP_R3_1.CheckTimer) ,XIO(MC_SP_R3_1.CW.[CWD.FAULT]) OTU(MC_SP_R3_1.CW.[CWD.FAULTLOGGED]) ,[GEQ(MC_SP_R3_1.CheckTimer,MC_SP_R3_1.CheckTime) [XIC(MC_SP_R3_1.CW.[CWD.OUTPUT]) XIO(MC_SP_R3_1.CW.[CWD.RUNFB]) ,XIO(MC_SP_R3_1.CW.[CWD.OUTPUT]) XIC(MC_SP_R3_1.CW.[CWD.RUNFB]) ] ,XIO(MC_SP_R3_1.CW.[CWD.HEALTHYFB]) ,XIO(MC_SP_R3_1.CW.[CWD.NOTTRIPPEDFB]) ,XIC(MC_SP_R3_1.CW.[CWD.FAULT]) XIC(Item_Faults_Are_Latched) ,XIC(MC_SP_R3_1.CW.[CWD.HIGHLIGHT]) ] XIO(MC_SP_R3_1.CW.[CWD.CHECKOFF]) XIO(Alarm_Reset) [OTE(MC_SP_R3_1.CW.[CWD.FAULT]) ,ALMD(MC_SP_R3_1_ALARM,0,0,0,0) ] ,XIC(MC_SP_R3_1.CW.[CWD.OUTPUT]) OTE(MC_SP_R3_1.CW.[CWD.PREVSCAN]) ,XIC(MC_SP_R3_1.CW.[CWD.FAULT]) EQU(Scada_Pump_Fault_No,0) XIO(MC_SP_R3_1.CW.[CWD.FAULTLOGGED]) [MOV(20001,Scada_Pump_Fault_No) ,OTL(MC_SP_R3_1.CW.[CWD.FAULTLOGGED]) ] ,XIO(MC_SP_R3_1.CW.[CWD.HEALTHYFB]) EQU(Scada_Pump_H_Fault_No,0) XIO(MC_SP_R3_1.CW.[CWD.HEALTHYFAULTLOGGED]) [MOV(20001,Scada_Pump_H_Fault_No) ,OTL(MC_SP_R3_1.CW.[CWD.HEALTHYFAULTLOGGED]) ] ,XIO(MC_SP_R3_1.CW.[CWD.NOTTRIPPEDFB]) EQU(Scada_Pump_H_Fault_No,0) XIO(MC_SP_R3_1.CW.[CWD.TRIPPEDFAULTLOGGED]) [MOV(20001,Scada_Pump_T_Fault_No) ,OTL(MC_SP_R3_1.CW.[CWD.TRIPPEDFAULTLOGGED]) ] ];